// TIA Portal project "EEEB EMBU 4_V17" (V17)

(* hardware
DEVICE "ET 200SP station_1"  ET 200SP-Station
   slot 0: "Rack_0"  Rack  6ES5 710-8MAx1
   slot 1: "EEEB EMBU"  CPU 1510SP-1 PN  6ES7 510-1DJ01-0AB0  V2.6
   slot 2: "SLOT1"  DI 16x24VDC ST  6ES7 131-6BH01-0BA0  V0.0
      slot 1: "SLOT1"  DI 16x24VDC ST
   slot 3: "SLOT2"  DI 16x24VDC ST  6ES7 131-6BH01-0BA0  V0.0
      slot 1: "SLOT2"  DI 16x24VDC ST
   slot 4: "SLOT3"  DI 16x24VDC ST  6ES7 131-6BH01-0BA0  V0.0
      slot 1: "SLOT3"  DI 16x24VDC ST
   slot 5: "SLOT4"  DI 16x24VDC ST  6ES7 131-6BH01-0BA0  V0.0
      slot 1: "SLOT4"  DI 16x24VDC ST
   slot 6: "SLOT5"  DI 16x24VDC ST  6ES7 131-6BH01-0BA0  V0.0
      slot 1: "SLOT5"  DI 16x24VDC ST
   slot 7: "SLOT6"  DQ 16x24VDC/0.5A ST  6ES7 132-6BH01-0BA0  V0.0
      slot 1: "SLOT6"  DQ 16x24VDC/0.5A ST
   slot 8: "SLOT7"  DQ 16x24VDC/0.5A ST  6ES7 132-6BH01-0BA0  V0.0
      slot 1: "SLOT7"  DQ 16x24VDC/0.5A ST
   slot 9: "SLOT8"  AI 8xI 2-,4-wire BA  6ES7 134-6GF00-0AA1  V1.0
      slot 1: "SLOT8"  AI 8xI 2-,4-wire BA
   slot 10: "SLO9"  AI 8xI 2-,4-wire BA  6ES7 134-6GF00-0AA1  V1.0
      slot 1: "SLO9"  AI 8xI 2-,4-wire BA
   slot 11: "SLOT10"  AQ 4xU/I ST  6ES7 135-6HD00-0BA1  V1.1
      slot 1: "SLOT10"  AQ 4xU/I ST
   slot 12: "SLOT11"  AQ 4xU/I ST  6ES7 135-6HD00-0BA1  V1.1
      slot 1: "SLOT11"  AQ 4xU/I ST
   slot 13: "Server module_1"  Server module  6ES7 193-6PA00-0AA0  V1.1
      slot 1: "Server module_1"  Server module
   slot 127: "BA 2xRJ45"  BA 2xRJ45  6ES7 193-6AR00-0AA0  V0.0
      slot 32769: "Port_1"  6ES7 193-6AR00-0AA0
      slot 32770: "Port_2"  6ES7 193-6AR00-0AA0
DEVICE "HMI_1"  KTP700 Basic PN
   slot 0: "HMI_1"  KTP700 Basic PN  6AV2 123-2GB03-0AX0  15.1.0.0
   slot 1: "HMI_RT_1"  KTP700 Basic PN  6AV2 123-2GB03-0AX0  15.1.0.0
   slot 5: "HMI_1.IE_CP_1"  PROFINET Interface  15.0.1.0
      slot 1: "PROFINET Interface_1"  PROFINET Interface
         slot 1: "Port_1"  Port
*)

// ===== PLC "EEEB EMBU"  CPU 1510SP-1 PN =====

VAR_GLOBAL   // PLC tag table "Default tag table"
   "System_Byte" AT %MB1 : Byte;
   "FirstScan" AT %M1.0 : Bool;
   "DiagStatusUpdate" AT %M1.1 : Bool;
   "AlwaysTRUE" AT %M1.2 : Bool;
   "AlwaysFALSE" AT %M1.3 : Bool;
   "Clock_Byte" AT %MB0 : Byte;
   "Clock_10Hz" AT %M0.0 : Bool;
   "Clock_5Hz" AT %M0.1 : Bool;
   "Clock_2.5Hz" AT %M0.2 : Bool;
   "Clock_2Hz" AT %M0.3 : Bool;
   "Clock_1.25Hz" AT %M0.4 : Bool;
   "Clock_1Hz" AT %M0.5 : Bool;
   "Clock_0.625Hz" AT %M0.6 : Bool;
   "Clock_0.5Hz" AT %M0.7 : Bool;
   "Tag_3" AT %M50.0 : Bool;
   "bloqueio_provisorio" AT %M2.0 : Bool;
   "pause" AT %M2.1 : Bool;
   "bloqueio_provisorio_1" AT %M2.2 : Bool;
   "Tag_4" AT %M83.0 : Bool;
   "CON_MOD" AT %MW80 : Int;
   "INI" AT %M82.0 : Bool;
END_VAR

VAR_GLOBAL   // PLC tag table "IO"
   "PCM_EEE_EMER" AT %I0.0 : Bool;   // PCM-E-CF-01-04 BOTAO DE EMERGENCIA - ATUADO
   "PCM_EEE_K27" AT %I0.1 : Bool;   // PCM-E-CF-01-04 RELE DE PROTECAO FUNCAO 27 - ATUADO
   "PCM_EEE_DJL" AT %I0.2 : Bool;   // PCM-E-CF-01-04 DISJUNTOR GERAL STATUS - LIGADO
   "PCM_EEE_DJD" AT %I0.3 : Bool;   // PCM-E-CF-01-04 DISJUNTOR GERAL STATUS - DESLIGADO
   "PCM_EEE_DJYFAL" AT %I0.4 : Bool;   // PCM-E-CF-01-04 DISJUNTOR GERAL STATUS - FALHA
   "PCM_EEE_DJFG" AT %I0.5 : Bool;   // PCM-E-CF-01-04 FALHA GERAL ATUADO
   "PCM_EEE_TR01_KA3" AT %I0.6 : Bool;   // PCM-E-CF-01-04 TRANSFORMADOR -TR-01 ALARME TEMP 150°
   "PCM_EEE_TR01_KA4" AT %I0.7 : Bool;   // PCM-E-CF-01-04 TRANSFORMADOR -TR-01 ALARME TEMP 155°
   "PCM_EEE_TR01_KA5" AT %I1.0 : Bool;   // PCM-E-CF-01-04 TRANSFORMADOR -TR-01 FALHA PROTECAO
   "PCM_EEE_INTRU" AT %I1.1 : Bool;   // PCM-E-CF-01-04 INTRUSAO NO PAINEL (COLUNA 01~04)
   "MB_01_FF" AT %I1.2 : Bool;   // MB-01 FALTA DE FASE
   "MB_01_MMNT" AT %I1.3 : Bool;   // MB-01 MODO MANUTENCAO
   "MB_01_ML" AT %I1.4 : Bool;   // MB-01 MODO LOCAL
   "MB_01_MA" AT %I1.5 : Bool;   // MB-01 MODO AUTOMATICO
   "MB_01_MN" AT %I1.6 : Bool;   // MB-01 MODO NORMAL
   "MB_01_HMNT" AT %I1.7 : Bool;   // MB-01 HABILITA MANUTENCAO
   "MB_01_BL" AT %I2.0 : Bool;   // MB-01 BOMBA LIGADA
   "MB_01_DINV" AT %I2.1 : Bool;   // MB-01 DEFEITO NO INVERSOR
   "MB_01_DMB" AT %I2.2 : Bool;   // MB-01 DEFEITO NA BOMBA
   "MB_01_RST" AT %I2.3 : Bool;   // MB-01 RESET
   "MB_01_INTRU" AT %I2.4 : Bool;   // MB-01 INTRUSAO NO PAINEL
   "MB_01_EMER" AT %I2.5 : Bool;   // MB-01 EMERGENCIA
   "MB_02_FF" AT %I2.6 : Bool;   // MB-02 FALTA DE FASE
   "MB_02_MMNT" AT %I2.7 : Bool;   // MB-02 MODO MANUTENCAO
   "MB_02_ML" AT %I3.0 : Bool;   // MB-02 MODO LOCAL
   "MB_02_MA" AT %I3.1 : Bool;   // MB-02 MODO AUTOMATICO
   "MB_02_MN" AT %I3.2 : Bool;   // MB-02 MODO NORMAL
   "MB_02_HMNT" AT %I3.3 : Bool;   // MB-02 HABILITA MANUTENCAO
   "MB_02_BL" AT %I3.4 : Bool;   // MB-02 BOMBA LIGADA
   "MB_02_DINV" AT %I3.5 : Bool;   // MB-02 DEFEITO NO INVERSOR
   "MB_02_DMB" AT %I3.6 : Bool;   // MB-02 DEFEITO NA BOMBA
   "MB_02_RST" AT %I3.7 : Bool;   // MB-02 RESET
   "MB_02_INTRU" AT %I4.0 : Bool;   // MB-02 INTRUSAO NO PAINEL
   "MB_02_EMER" AT %I4.1 : Bool;   // MB-02 EMERGENCIA
   "MB_03_FF" AT %I4.2 : Bool;   // MB-03 FALTA DE FASE
   "MB_03_MMNT" AT %I4.3 : Bool;   // MB-03 MODO MANUTENCAO
   "MB_03_ML" AT %I4.4 : Bool;   // MB-03 MODO LOCAL
   "MB_03_MA" AT %I4.5 : Bool;   // MB-03 MODO AUTOMATICO
   "MB_03_MN" AT %I4.6 : Bool;   // MB-03 MODO NORMAL
   "MB_03_HMNT" AT %I4.7 : Bool;   // MB-03 HABILITA MANUTENCAO
   "MB_03_BL" AT %I5.0 : Bool;   // MB-03 BOMBA LIGADA
   "MB_03_DINV" AT %I5.1 : Bool;   // MB-03 DEFEITO NO INVERSOR
   "MB_03_DMB" AT %I5.2 : Bool;   // MB-03 DEFEITO NA BOMBA
   "MB_03_RST" AT %I5.3 : Bool;   // MB-03 RESET
   "MB_03_INTRU" AT %I5.4 : Bool;   // MB-03 INTRUSAO NO PAINEL
   "MB_03_EMER" AT %I5.5 : Bool;   // MB-03EMERGENCIA
   "MB_04_FF" AT %I5.6 : Bool;   // MB-04 FALTA DE FASE
   "MB_04_MMNT" AT %I5.7 : Bool;   // MB-04 MODO MANUTENCAO
   "MB_04_ML" AT %I6.0 : Bool;   // MB-04 MODO LOCAL
   "MB_04_MA" AT %I6.1 : Bool;   // MB-04 MODO AUTOMATICO
   "MB_04_MN" AT %I6.2 : Bool;   // MB-04 MODO NORMAL
   "MB_04_HMNT" AT %I6.3 : Bool;   // MB-04 HABILITA MANUTENCAO
   "MB_04_BL" AT %I6.4 : Bool;   // MB-04 BOMBA LIGADA
   "MB_04_DINV" AT %I6.5 : Bool;   // MB-04 DEFEITO NO INVERSOR
   "MB_04_DMB" AT %I6.6 : Bool;   // MB-04 DEFEITO NA BOMBA
   "MB_04_RST" AT %I6.7 : Bool;   // MB-04 RESET
   "MB_04_INTRU" AT %I7.0 : Bool;   // MB-04 INTRUSAO NO PAINEL
   "MB_04_EMER" AT %I7.1 : Bool;   // MB-04 EMERGENCIA
   "QGBT_EMER" AT %I7.2 : Bool;   // QGBT-AUX-01 BOTAO DE EMERGENCIA ATUADO
   "QGBT_K27" AT %I7.3 : Bool;   // QGBT-AUX-01 RELE DE PROTECAO FUNCAO 27/59 ATUADO
   "QGBT_DISJ_LIG" AT %I7.4 : Bool;   // QGBT-AUX-01 DISJUNTOR GERAL STATUS - LIGADO
   "QGBT_DISJ_DESLIG" AT %I7.5 : Bool;   // QGBT-AUX-01 DISJUNTOR GERAL STATUS - DESLIGADO
   "QGBT_DISJ_YFAL" AT %I7.6 : Bool;   // QGBT-AUX-01 DISJUNTOR GERAL FALHA - TRIP
   "QGBT_INTRU" AT %I7.7 : Bool;   // QGBT-AUX-01 INTRUSAO NO PAINEL
   "KI165" AT %I8.0 : Bool;   // RESERVA
   "KI166" AT %I8.1 : Bool;   // RESERVA
   "KI167" AT %I8.2 : Bool;   // RESERVA
   "KI168" AT %I8.3 : Bool;   // RESERVA
   "KI169" AT %I8.4 : Bool;   // RESERVA
   "KI170" AT %I8.5 : Bool;   // RESERVA
   "KI171" AT %I8.6 : Bool;   // RESERVA
   "KI172" AT %I8.7 : Bool;   // RESERVA
   "LSL_001" AT %I9.0 : Bool;   // CHAVE DE NIVEL -LSL-001
   "LSH_001" AT %I9.1 : Bool;   // CHAVE DE NIVEL -LSH-001
   "LSL_002" AT %I9.2 : Bool;   // CHAVE DE NIVEL -LSL-002
   "LSH_002" AT %I9.3 : Bool;   // CHAVE DE NIVEL -LSH-002
   "PCE_EEE_INTRU" AT %I9.4 : Bool;   // INTRUSAO NO PAINEL
   "PCE_EEE_UPS_ALM" AT %I9.5 : Bool;   // UPS EM ALARME FALHA NA BATERIA
   "PCE_EEE_UPS_FE" AT %I9.6 : Bool;   // UPS EM OPERACAO FALTA DE ENERGIA
   "PCE_EEE_UPS_CHAR" AT %I9.7 : Bool;   // UPS EM ALARME BATERIA CARREGADA
   "MB_01_SH" AT %Q0.0 : Bool;   // MB-01 SOLICITACAO HIDRAULICA
   "MB_01_PH" AT %Q0.1 : Bool;   // MB-01 PROTECAO HIDRAULICA
   "MB_01_INTV" AT %Q0.2 : Bool;   // MB-01 INTERVALO (COM)
   "MB_01_RR" AT %Q0.3 : Bool;   // MB-01 RESET REMOTO
   "MB_01_INTVS" AT %Q0.4 : Bool;   // MB-01 INTERVALO SINAL
   "MB_02_SH" AT %Q0.5 : Bool;   // MB-02 SOLICITACAO HIDRAULICA
   "MB_02_PH" AT %Q0.6 : Bool;   // MB-02 PROTECAO HIDRAULICA
   "MB_02_INTV" AT %Q0.7 : Bool;   // MB-02 INTERVALO (COM)
   "MB_02_RR" AT %Q1.0 : Bool;   // MB-02 RESET REMOTO
   "MB_02_INTVS" AT %Q1.1 : Bool;   // MB-02 INTERVALO SINAL
   "MB_03_SH" AT %Q1.2 : Bool;   // MB-03 SOLICITACAO HIDRAULICA
   "MB_03_PH" AT %Q1.3 : Bool;   // MB-03 PROTECAO HIDRAULICA
   "MB_03_INTV" AT %Q1.4 : Bool;   // MB-03 INTERVALO (COM)
   "MB_03_RR" AT %Q1.5 : Bool;   // MB-03 RESET REMOTO
   "MB_03_INTVS" AT %Q1.6 : Bool;   // MB-03 INTERVALO SINAL
   "MB_04_SH" AT %Q1.7 : Bool;   // MB-04 SOLICITACAO HIDRAULICA
   "LIT_001" AT %IW10 : Int;   // -LIT-001 TRANSMISSOR DE NIVEL TANQUE (TIPO RADAR)
   "MB_01_REF_VEL" AT %IW12 : Int;   // REFERENCIA DE VELOCIDADE INVERSOR DE FREQUENCIA BOMBA 01
   "MB_02_REF_VEL" AT %IW14 : Int;   // REFERENCIA DE VELOCIDADE INVERSOR DE FREQUENCIA BOMBA 02
   "MB_03_REF_VEL" AT %IW16 : Int;   // REFERENCIA DE VELOCIDADE INVERSOR DE FREQUENCIA BOMBA 03
   "MB_04_REF_VEL" AT %IW18 : Int;   // REFERENCIA DE VELOCIDADE INVERSOR DE FREQUENCIA BOMBA 04
   "FB6" AT %IW20 : Int;   // RESERVA
   "FB7" AT %IW22 : Int;   // RESERVA
   "FB8" AT %IW24 : Int;   // RESERVA
   "FB9" AT %IW26 : Int;   // RESERVA
   "FB10" AT %IW28 : Int;   // RESERVA
   "FB11" AT %IW30 : Int;   // RESERVA
   "FB12" AT %IW32 : Int;   // RESERVA
   "FB13" AT %IW34 : Int;   // RESERVA
   "FB14" AT %IW36 : Int;   // RESERVA
   "FB15" AT %IW38 : Int;   // RESERVA
   "FB16" AT %IW40 : Int;   // RESERVA
   "MB_01_VEL" AT %QW4 : Int;   // SETPOINT INVERSOR DE FREQUENCIA BOMBA 01
   "MB_02_VEL" AT %QW6 : Int;   // SETPOINT INVERSOR DE FREQUENCIA BOMBA 02
   "MB_03_VEL" AT %QW8 : Int;   // SETPOINT INVERSOR DE FREQUENCIA BOMBA 03
   "MB_04_VEL" AT %QW10 : Int;   // SETPOINT INVERSOR DE FREQUENCIA BOMBA 04
   "F25" AT %QW12 : Int;   // RESERVA
   "F26" AT %QW14 : Int;   // RESERVA
   "F27" AT %QW16 : Int;   // RESERVA
   "F28" AT %QW18 : Int;   // RESERVA
   "MB_04_PH" AT %Q2.0 : Bool;   // MB-04 PROTECAO HIDRAULICA
   "MB_04_INTV" AT %Q2.1 : Bool;   // MB-04 INTERVALO (COM)
   "MB_04_RR" AT %Q2.2 : Bool;   // MB-04 RESET REMOTO
   "MB_04_INTVS" AT %Q2.3 : Bool;   // MB-04 INTERVALO SINAL
   "KO21" AT %Q2.4 : Bool;   // RESERVA
   "KO22" AT %Q2.5 : Bool;   // RESERVA
   "KO23" AT %Q2.6 : Bool;   // RESERVA
   "KO24" AT %Q2.7 : Bool;   // RESERVA
   "KO25" AT %Q3.0 : Bool;   // RESERVA
   "KO26" AT %Q3.1 : Bool;   // RESERVA
   "KO27" AT %Q3.2 : Bool;   // RESERVA
   "KO28" AT %Q3.3 : Bool;   // RESERVA
   "KO29" AT %Q3.4 : Bool;   // RESERVA
   "KO30" AT %Q3.5 : Bool;   // RESERVA
   "KO31" AT %Q3.6 : Bool;   // RESERVA
   "KO32" AT %Q3.7 : Bool;   // RESERVA
END_VAR

VAR_GLOBAL   // PLC tag table "ALARMES"
   "ALM0" AT %MW100 : Word;   // ALARMES MB-01
   "ALM2" AT %MW102 : Word;   // ALARMES MB-02
   "ALM4" AT %MW104 : Word;   // ALARMES MB-03
   "ALM6" AT %MW106 : Word;   // ALARMES MB-04
   "ALM8" AT %MW108 : Word;   // ALARMES LIT_001
   "ALM10" AT %MW110 : Word;   // ALARMES PCM-EEE
   "ALM12" AT %MW112 : Word;   // ALARMES QGBT
   "ALM14" AT %MW114 : Word;   // ALARMES CHAVE DE NIVEL
   "ALM16" AT %MW116 : Word;   // ALARMES PCE-EEE
END_VAR

DATA_BLOCK "DIVERSOS"   // DB1
{ S7_Optimized_Access := 'TRUE' }
VERSION : 0.1
   VAR
      T1S : Bool;   // PULSO A CADA 1 SEGUNDO
      AUX_T1S : Bool;   // PULSO A CADA 1 SEGUNDO
      QTDE_PULSO : DInt := 200;
      ForcePulso : Bool;
      N_L00P : Int;
      Aux_N_LOOP : Int;
      Looping : Int := 0;
      TMR : Array[0..10] of IEC_TIMER;
      P1S : Bool;   // Pulso de 1 segundo
      "MB-01-SP" : Bool;   // Solicitação partida de bomba
      "MB-02-SP" : Bool;   // Solicitação partida de bomba
      "MB-03-SP" : Bool;   // Solicitação partida de bomba
      "MB-04-SP" : Bool;   // Solicitação partida de bomba
   END_VAR
BEGIN
END_DATA_BLOCK

DATA_BLOCK "INTPRO_DB"   // DB2
{ S7_Optimized_Access := 'TRUE' }
VERSION : 0.1
// stored: InstanceOfName INTPRO
"INTPRO"
BEGIN
END_DATA_BLOCK

DATA_BLOCK "LOOP_DB"   // DB3
{ S7_Optimized_Access := 'TRUE' }
VERSION : 0.1
// stored: InstanceOfName LOOP
"LOOP"
BEGIN
END_DATA_BLOCK

DATA_BLOCK "ROD4_DB"   // DB9
{ S7_Optimized_Access := 'FALSE' }
VERSION : 0.1
// stored: InstanceOfName ROD4
"ROD4"
BEGIN
END_DATA_BLOCK

DATA_BLOCK "ANALOGICOS_DB"   // DB101
{ S7_Optimized_Access := 'TRUE' }
VERSION : 0.1
// stored: InstanceOfName ANALOGICOS
"ANALOGICOS"
BEGIN
END_DATA_BLOCK

DATA_BLOCK "MODBUS_DB"   // DB102
{ S7_Optimized_Access := 'TRUE' }
VERSION : 0.1
// stored: InstanceOfName MODBUS
"MODBUS"
BEGIN
END_DATA_BLOCK

DATA_BLOCK "Digitais"   // DB300
{ S7_Optimized_Access := 'FALSE' }
VERSION : 0.1
   VAR
      "MB-01-YSH" : Bool;   // Elevatoria principal 1 ligado
      "MB-01-YR" : Bool;   // Elevatoria principal 1 remoto
      "MB-01-YF" : Bool;   // Elevatoria principal 1 falha
      "MB-01-YFF" : Bool;   // Elevatoria principal 1 falta de fase
      "MB-01-MM" : Bool;   // Elevatoria principal 1 modo manutenção
      "MB-01-MA" : Bool;   // Elevatoria principal 1 modo automatico
      "MB-01-EMER" : Bool;   // Elevatoria principal 1 emergencia
      "MB-01-MN" : Bool;   // Elevatoria principal 1 modo normal
      "MB-01-ML" : Bool;   // Elevatoria principal 1 modo local
      "MB-01-YFI" : Bool;   // Elevatoria principal 1 com falha no inversor
      "MB-01-YFA" : Bool;   // Elevatoria principal 1 com falha no acionamento
      "MB-01-YPTA" : Bool;   // Elevatoria principal 1 com proteção térmica atuada
      "MB-01-HM" : Bool;   // Elevatoria principal 1 habilita manutenção
      "MB-01-RST" : Bool;   // Elevatoria principal 1 reset
      "MB-01-INTRU" : Bool;   // Elevatoria principal 1 intrusão no painel
      "MB-01-YFB" : Bool;   // Elevatoria principal 1 defeito na bomba
      "MB-02-YSH" : Bool;   // Elevatoria principal 2 ligado
      "MB-02-YR" : Bool;   // Elevatoria principal 2 remoto
      "MB-02-YF" : Bool;   // Elevatoria principal 2 falha
      "MB-02-YFF" : Bool;   // Elevatoria principal 2 falta de fase
      "MB-02-MM" : Bool;   // Elevatoria principal 2 modo manutenção
      "MB-02-MA" : Bool;   // Elevatoria principal 2 modo automatico
      "MB-02-EMER" : Bool;   // Elevatoria principal 2 emergencia
      "MB-02-MN" : Bool;   // Elevatoria principal 2 modo normal
      "MB-02-ML" : Bool;   // Elevatoria principal 2 modo local
      "MB-02-YFI" : Bool;   // Elevatoria principal 2 com falha no inversor
      "MB-02-YFA" : Bool;   // Elevatoria principal 2 com falha no acionamento
      "MB-02-YPTA" : Bool;   // Elevatoria principal 2 com proteção térmica atuada
      "MB-02-HM" : Bool;   // Elevatoria principal 2 habilita manutenção
      "MB-02-RST" : Bool;   // Elevatoria principal 2 reset
      "MB-02-INTRU" : Bool;   // Elevatoria principal 2 intrusão no painel
      "MB-02-YFB" : Bool;   // Elevatoria principal 2 defeito na bomba
      "MB-03-YSH" : Bool;   // Elevatoria principal 3 ligado
      "MB-03-YR" : Bool;   // Elevatoria principal 3 remoto
      "MB-03-YF" : Bool;   // Elevatoria principal 3 falha
      "MB-03-YFF" : Bool;   // Elevatoria principal 3 falta de fase
      "MB-03-MM" : Bool;   // Elevatoria principal 3 modo manutenção
      "MB-03-MA" : Bool;   // Elevatoria principal 3 modo automatico
      "MB-03-EMER" : Bool;   // Elevatoria principal 3 emergencia
      "MB-03-MN" : Bool;   // Elevatoria principal 3 modo normal
      "MB-03-ML" : Bool;   // Elevatoria principal 3 modo local
      "MB-03-YFI" : Bool;   // Elevatoria principal 3 com falha no inversor
      "MB-03-YFA" : Bool;   // Elevatoria principal 3 com falha no acionamento
      "MB-03-YPTA" : Bool;   // Elevatoria principal 3 com proteção térmica atuada
      "MB-03-HM" : Bool;   // Elevatoria principal 3 habilita manutenção
      "MB-03-RST" : Bool;   // Elevatoria principal 3 reset
      "MB-03-INTRU" : Bool;   // Elevatoria principal 3 intrusão no painel
      "MB-03-YFB" : Bool;   // Elevatoria principal 3 defeito na bomba
      "MB-04-YSH" : Bool;   // Elevatoria principal 4 ligado
      "MB-04-YR" : Bool;   // Elevatoria principal 4 remoto
      "MB-04-YF" : Bool;   // Elevatoria principal 4 falha
      "MB-04-YFF" : Bool;   // Elevatoria principal 4 falta de fase
      "MB-04-MM" : Bool;   // Elevatoria principal 4 modo manutenção
      "MB-04-MA" : Bool;   // Elevatoria principal 4 modo automatico
      "MB-04-EMER" : Bool;   // Elevatoria principal 4 emergencia
      "MB-04-MN" : Bool;   // Elevatoria principal 4 modo normal
      "MB-04-ML" : Bool;   // Elevatoria principal 4 modo local
      "MB-04-YFI" : Bool;   // Elevatoria principal 4 com falha no inversor
      "MB-04-YFA" : Bool;   // Elevatoria principal 4 com falha no acionamento
      "MB-04-YPTA" : Bool;   // Elevatoria principal 4 com proteção térmica atuada
      "MB-04-HM" : Bool;   // Elevatoria principal 4 habilita manutenção
      "MB-04-RST" : Bool;   // Elevatoria principal 4 reset
      "MB-04-INTRU" : Bool;   // Elevatoria principal 4 intrusão no painel
      "MB-04-YFB" : Bool;   // Elevatoria principal 4 defeito na bomba
      "LIT_001-AL8" : Bool;   // Disponível para alarme
      "LIT_001-AL9" : Bool;   // Disponível para alarme
      "LIT_001-AL10" : Bool;   // Disponível para alarme
      "LIT_001-AL11" : Bool;   // Disponível para alarme
      "LIT_001-AL12" : Bool;   // Disponível para alarme
      "LIT_001-AL13" : Bool;   // Disponível para alarme
      "LIT_001-AL14" : Bool;   // Disponível para alarme
      "LIT_001-AL15" : Bool;   // Disponível para alarme
      "LIT_001-YHH" : Bool;   // Alarme de nível muito alto do tanque
      "LIT_001-YH" : Bool;   // Alarme de nível alto do tanque
      "LIT_001-YL" : Bool;   // Alarme de nível baixo do tanque
      "LIT_001-YLL" : Bool;   // Alarme de nível muito baixo do tanque
      "LIT_001-YFS" : Bool;   // Transmissor de nível do tanque com falha de sinal
      "LIT_001-AL5" : Bool;   // Disponível para alarme
      "LIT_001-AL6" : Bool;   // Disponível para alarme
      "LIT_001-AL7" : Bool;   // Disponível para alarme
      PCM_EEE_EMER : Bool;   // PCM-E-CF-01-04 BOTAO DE EMERGENCIA - ATUADO
      PCM_EEE_K27 : Bool;   // PCM-E-CF-01-04 RELE DE PROTECAO FUNCAO 27 - ATUADO
      PCM_EEE_DISJ_LIG : Bool;   // PCM-E-CF-01-04 DISJUNTOR GERAL STATUS - LIGADO
      PCM_EEE_DISJ_DESLIG : Bool;   // PCM-E-CF-01-04 DISJUNTOR GERAL STATUS - DESLIGADO
      PCM_EEE_DISJ_YFAL : Bool;   // PCM-E-CF-01-04 DISJUNTOR GERAL STATUS - FALHA
      PCM_EEE_DISJ_FAL_GR : Bool;   // PCM-E-CF-01-04 FALHA GERAL ATUADO
      PCM_EEE_TR01_KA3 : Bool;   // PCM-E-CF-01-04 TRANSFORMADOR -TR-01 ALARME TEMP 150°
      PCM_EEE_TR01_KA4 : Bool;   // PCM-E-CF-01-04 TRANSFORMADOR -TR-01 ALARME TEMP 155°
      PCM_EEE_TR01_KA5 : Bool;   // PCM-E-CF-01-04 TRANSFORMADOR -TR-01 FALHA PROTECAO
      PCM_EEE_INTRU : Bool;   // PCM-E-CF-01-04 INTRUSAO NO PAINEL (COLUNA 01~04)
      PCM_EEE_RSERVA_0 : Bool;   // PCM-E-CF-01-04 BIT RESERVA DA WORD
      PCM_EEE_RSERVA_1 : Bool;   // PCM-E-CF-01-04 BIT RESERVA DA WORD
      PCM_EEE_RSERVA_2 : Bool;   // PCM-E-CF-01-04 BIT RESERVA DA WORD
      PCM_EEE_RSERVA_3 : Bool;   // PCM-E-CF-01-04 BIT RESERVA DA WORD
      PCM_EEE_RSERVA_4 : Bool;   // PCM-E-CF-01-04 BIT RESERVA DA WORD
      PCM_EEE_RSERVA_5 : Bool;   // PCM-E-CF-01-04 BIT RESERVA DA WORD
      QGBT_EMER : Bool;   // QGBT-AUX-01 BOTAO DE EMERGENCIA ATUADO
      QGBT_K27 : Bool;   // QGBT-AUX-01 RELE DE PROTECAO FUNCAO 27/59 ATUADO
      QGBT_DJL : Bool;   // QGBT-AUX-01 DISJUNTOR GERAL STATUS - LIGADO
      QGBT_DJD : Bool;   // QGBT-AUX-01 DISJUNTOR GERAL STATUS - DESLIGADO
      QGBT_DJYFAL : Bool;   // QGBT-AUX-01 DISJUNTOR GERAL FALHA - TRIP
      QGBT_INTRU : Bool;   // QGBT-AUX-01 INTRUSAO NO PAINEL
      QGBT_RESERVA_0 : Bool;   // QGBT-AUX-01 BIT RESERVA DA WORD
      QGBT_RESERVA_1 : Bool;   // QGBT-AUX-01 BIT RESERVA DA WORD
      QGBT_RESERVA_2 : Bool;   // QGBT-AUX-01 BIT RESERVA DA WORD
      QGBT_RESERVA_3 : Bool;   // QGBT-AUX-01 BIT RESERVA DA WORD
      QGBT_RESERVA_4 : Bool;   // QGBT-AUX-01 BIT RESERVA DA WORD
      QGBT_RESERVA_5 : Bool;   // QGBT-AUX-01 BIT RESERVA DA WORD
      QGBT_RESERVA_6 : Bool;   // QGBT-AUX-01 BIT RESERVA DA WORD
      QGBT_RESERVA_7 : Bool;   // QGBT-AUX-01 BIT RESERVA DA WORD
      QGBT_RESERVA_8 : Bool;   // QGBT-AUX-01 BIT RESERVA DA WORD
      QGBT_RESERVA_9 : Bool;   // QGBT-AUX-01 BIT RESERVA DA WORD
      LSL_001 : Bool;   // CHAVE DE NIVEL -LSL-001
      LSH_001 : Bool;   // CHAVE DE NIVEL -LSH-001
      LSL_002 : Bool;   // CHAVE DE NIVEL -LSL-002
      LSH_002 : Bool;   // CHAVE DE NIVEL -LSH-002
      LS_RESERVA_0 : Bool;   // CHAVE DE NIVEL - LS BIT RESERVA DA WORD
      LS_RESERVA_1 : Bool;   // CHAVE DE NIVEL - LS BIT RESERVA DA WORD
      LS_RESERVA_2 : Bool;   // CHAVE DE NIVEL - LS BIT RESERVA DA WORD
      LS_RESERVA_3 : Bool;   // CHAVE DE NIVEL - LS BIT RESERVA DA WORD
      LS_RESERVA_4 : Bool;   // CHAVE DE NIVEL - LS BIT RESERVA DA WORD
      LS_RESERVA_5 : Bool;   // CHAVE DE NIVEL - LS BIT RESERVA DA WORD
      LS_RESERVA_6 : Bool;   // CHAVE DE NIVEL - LS BIT RESERVA DA WORD
      LS_RESERVA_7 : Bool;   // CHAVE DE NIVEL - LS BIT RESERVA DA WORD
      LS_RESERVA_8 : Bool;   // CHAVE DE NIVEL - LS BIT RESERVA DA WORD
      LS_RESERVA_9 : Bool;   // CHAVE DE NIVEL - LS BIT RESERVA DA WORD
      LS_RESERVA_10 : Bool;   // CHAVE DE NIVEL - LS BIT RESERVA DA WORD
      LS_RESERVA_11 : Bool;   // CHAVE DE NIVEL - LS BIT RESERVA DA WORD
      PCE_EEE_INTRU : Bool;   // INTRUSAO NO PAINEL
      PCE_EEE_UPS_ALM : Bool;   // UPS EM ALARME FALHA NA BATERIA
      PCE_EEE_UPS_FE : Bool;   // UPS EM OPERACAO FALTA DE ENERGIA
      PCE_EEE_UPS_CHAR : Bool;   // UPS EM ALARME BATERIA CARREGADA
      "PCM-E-CF-01-P100-YFC" : Bool;   // Falha de comunicação com medidor do PCM-E-CF-01
      "QGBT-AUX-01-P100-YFC" : Bool;   // Falha de comunicação com medidor do PCM-E-CF-02
   END_VAR
BEGIN
END_DATA_BLOCK

DATA_BLOCK "ALARMES"   // DB301
{ S7_Optimized_Access := 'TRUE' }
VERSION : 0.1
   VAR
      "CCM-02-EA-P100-YFC" : Bool;   // Falha de comunicação com medidor do CCM1
      "CCM-02-EB-P100-YFC" : Bool;   // Falha de comunicação com medidor do CCM2
      "LIT_001-YHH" : Bool;   // Alarme de nível muito alto do tanque água bruta
      "LIT_001-YH" : Bool;   // Alarme de nível alto do tanque água bruta
      "LIT_001-YL" : Bool;   // Alarme de nível baixo do tanque água bruta
      "LIT_001-YLL" : Bool;   // Alarme de nível muito baixo do tanque água bruta
      "LIT_001-YFS" : Bool;   // Transmissor de nível do tanque água bruta com falha de sinal
      "LIT_001-YHHH" : Bool;   // Alarme de nível muito alto - desliga CAB e lavagem peneira
      "CAB-PT-015-YH" : Bool;
      "CAB-PT-015-YFS" : Bool;
      "MB-03-YIP" : Bool;   // MB-03 com intervalo entre partidas
      "MB-02-YIP" : Bool;   // MB-02 com intervalo entre partidas
      "MB-01-YIP" : Bool;   // MB-01 com intervalo entre partidas
   END_VAR
BEGIN
END_DATA_BLOCK

DATA_BLOCK "STATUS"   // DB302
{ S7_Optimized_Access := 'FALSE' }
VERSION : 0.1
   VAR
      "SO-203-06A-YI" : Bool;   // Soprador tanque de aeração intertravado
      "SO-203-06B-YI" : Bool;   // Soprador tanque de aeração intertravado
      "SO-203-06C-YI" : Bool;   // Soprador tanque de aeração intertravado
      "SO-203-06D-YI" : Bool;   // Soprador tanque de aeração intertravado
      "SO-203-06E-YI" : Bool;   // Soprador tanque de aeração intertravado
      "SO-203-06F-YI" : Bool;   // Soprador tanque de aeração intertravado
      "MB-01-YSP" : Bool;   // MB-01 selecionada como principal
      "MB-02-YSP" : Bool;   // MB-02 selecionada como principal
      "MB-04-YSP" : Bool;   // MB-03 selecionada como principal
      "MB-03-YSP" : Bool;   // MB-03 selecionada como principal
      "MB-01-YC1" : Bool;   // MB-01 selecionada como complementar 1
      "MB-02-YC1" : Bool;   // MB-02 selecionada como complementar 1
      "MB-04-YC1" : Bool;   // MB-03 selecionada como complementar 1
      "MB-03-YC1" : Bool;   // MB-03 selecionada como complementar 1
      "MB-01-YC2" : Bool;   // MB-01 selecionada como complementar 2
      "MB-02-YC2" : Bool;   // MB-02 selecionada como complementar 2
      "MB-04-YC2" : Bool;   // MB-03 selecionada como complementar 2
      "MB-03-YC2" : Bool;   // MB-03 selecionada como complementar 2
      "MB-01-YC3" : Bool;   // MB-01 selecionada como complementar 3
      "MB-02-YC3" : Bool;   // MB-02 selecionada como complementar 3
      "MB-04-YC3" : Bool;   // MB-03 selecionada como complementar 3
      "MB-03-YC3" : Bool;   // MB-03 selecionada como complementar 3
   END_VAR
BEGIN
END_DATA_BLOCK

DATA_BLOCK "COMANDOS"   // DB303
{ S7_Optimized_Access := 'FALSE' }
VERSION : 0.1
   VAR
      "MB-01-HS9" : Bool := false;   // Comando disponível
      "MB-01-HS10" : Bool := false;   // Comando disponível
      "MB-01-HS11" : Bool;   // Comando disponível
      "MB-01-HS12" : Bool;   // Comando disponível
      "MB-01-HS13" : Bool;   // Comando disponível
      "MB-01-HS14" : Bool;   // Comando disponível
      "MB-01-HS15" : Bool;   // Comando disponível
      "MB-01-HS16" : Bool;   // Comando disponível
      "MB-01-HS1" : Bool := true;   // Comando manual/automático
      "MB-01-HS2" : Bool := false;   // Comando liga
      "MB-01-HS3" : Bool := false;   // Comando desliga
      "MB-01-HS4" : Bool := false;   // Comando reset falha
      "MB-01-HS5" : Bool := false;   // Comando reset tempo de operação
      "MB-01-HS6" : Bool;
      "MB-01-HS7" : Bool := false;   // Comando habilita bloqueio
      "MB-01-HS8" : Bool := false;   // Comando disponível
      "MB-02-HS9" : Bool := false;   // Comando disponível
      "MB-02-HS10" : Bool := false;   // Comando disponível
      "MB-02-HS11" : Bool;   // Comando disponível
      "MB-02-HS12" : Bool;   // Comando disponível
      "MB-02-HS13" : Bool;   // Comando disponível
      "MB-02-HS14" : Bool;   // Comando disponível
      "MB-02-HS15" : Bool;   // Comando disponível
      "MB-02-HS16" : Bool;   // Comando disponível
      "MB-02-HS1" : Bool := true;   // Comando manual/automático
      "MB-02-HS2" : Bool := false;   // Comando liga
      "MB-02-HS3" : Bool := false;   // Comando desliga
      "MB-02-HS4" : Bool := false;   // Comando reset falha
      "MB-02-HS5" : Bool := false;   // Comando reset tempo de operação
      "MB-02-HS6" : Bool;
      "MB-02-HS7" : Bool := false;   // Comando habilita bloqueio
      "MB-02-HS8" : Bool := false;   // Comando disponível
      "MB-03-HS9" : Bool := false;   // Comando disponível
      "MB-03-HS10" : Bool := false;   // Comando disponível
      "MB-03-HS11" : Bool;   // Comando disponível
      "MB-03-HS12" : Bool;   // Comando disponível
      "MB-03-HS13" : Bool;   // Comando disponível
      "MB-03-HS14" : Bool;   // Comando disponível
      "MB-03-HS15" : Bool;   // Comando disponível
      "MB-03-HS16" : Bool;   // Comando disponível
      "MB-03-HS1" : Bool := true;   // Comando manual/automático
      "MB-03-HS2" : Bool := false;   // Comando liga
      "MB-03-HS3" : Bool := false;   // Comando desliga
      "MB-03-HS4" : Bool := false;   // Comando reset falha
      "MB-03-HS5" : Bool := false;   // Comando reset tempo de operação
      "MB-03-HS6" : Bool;
      "MB-03-HS7" : Bool := false;   // Comando habilita bloqueio
      "MB-03-HS8" : Bool := false;   // Comando disponível
      "MB-04-HS9" : Bool := false;   // Comando disponível
      "MB-04-HS10" : Bool := false;   // Comando disponível
      "MB-04-HS11" : Bool;   // Comando disponível
      "MB-04-HS12" : Bool;   // Comando disponível
      "MB-04-HS13" : Bool;   // Comando disponível
      "MB-04-HS14" : Bool;   // Comando disponível
      "MB-04-HS15" : Bool;   // Comando disponível
      "MB-04-HS16" : Bool;   // Comando disponível
      "MB-04-HS1" : Bool := false;   // Comando manual/automático
      "MB-04-HS2" : Bool := false;   // Comando liga
      "MB-04-HS3" : Bool := false;   // Comando desliga
      "MB-04-HS4" : Bool := false;   // Comando reset falha
      "MB-04-HS5" : Bool := false;   // Comando reset tempo de operação
      "MB-04-HS6" : Bool;
      "MB-04-HS7" : Bool := false;   // Comando habilita bloqueio
      "MB-04-HS8" : Bool := false;   // Comando disponível
      "LIT_001-HS9" : Bool;   // Comando disponível
      "LIT_001-HS10" : Bool;   // Comando disponível
      "LIT_001-HS11" : Bool;   // Comando disponível
      "LIT_001-HS12" : Bool;   // Comando disponível
      "LIT_001-HS13" : Bool;   // Comando disponível
      "LIT_001-HS14" : Bool;   // Comando disponível
      "LIT_001-HS15" : Bool;   // Comando disponível
      "LIT_001-HS16" : Bool;   // Comando disponível
      "LIT_001-HSHH" : Bool;   // Inibe alarme muito alto montante peneira 1
      "LIT_001-HSH" : Bool;   // Inibe alarme nível alto montante peneira 1
      "LIT_001-HSL" : Bool;   // Inibe alarme nível baixo montante peneira 1
      "LIT_001-HSLL" : Bool;   // Inibe alarme nível muito baixo montante peneira 1
      "LIT_001-HSM" : Bool;   // Habilita valor manual para medidor
      "LIT_001-HS6" : Bool;   // Comando disponível
      "LIT_001-HS7" : Bool;   // Comando disponível
      "LIT_001-HS8" : Bool;   // Comando disponível
      "PID-TA3-HI" : Bool;   // Habilita integrall PID tanque de aeração
      "PID-EEEB-HD" : Bool;   // Habilita derivativo PID tanque de aeração
      "PID-EEEB-HP" : Bool;   // Habilita proporcional PID tanque de aeração
      "PID-EEEB-HI" : Bool;   // Habilita integrall PID tanque de aeração
      "PID-TA5-HD" : Bool;   // Habilita derivativo PID tanque de aeração
      "PID-TA5-HP" : Bool;   // Habilita proporcional PID tanque de aeração
      "PID-TA5-HI" : Bool;   // Habilita integrall PID tanque de aeração
      "PID-TA1-HM" : Bool;   // Habilita valor manual para saída
      "PID-TA1-HD" : Bool;   // Habilita derivativo PID tanque de aeração
      "PID-TA1-HP" : Bool;   // Habilita proporcional PID tanque de aeração
      "PID-TA1-HI" : Bool;   // Habilita integrall PID tanque de aeração
      "PID-TA2-HD" : Bool;   // Habilita derivativo PID tanque de aeração
      "PID-TA2-HP" : Bool;   // Habilita proporcional PID tanque de aeração
      "PID-TA2-HI" : Bool;   // Habilita integrall PID tanque de aeração
      "PID-TA3-HD" : Bool;   // Habilita derivativo PID tanque de aeração
      "PID-TA3-HP" : Bool;   // Habilita proporcional PID tanque de aeração
      "PID-TA2-HM" : Bool;   // Habilita valor manual para saída
      "PID-TA3-HM" : Bool;   // Habilita valor manual para saída
      "PID-EEEB-HM" : Bool;   // Habilita valor manual para saída
      "PID-TA5-HM" : Bool;   // Habilita valor manual para saída
   END_VAR
BEGIN
END_DATA_BLOCK

DATA_BLOCK "VARIAVEIS"   // DB304
{ S7_Optimized_Access := 'FALSE' }
VERSION : 0.1
   VAR
      "MB-01-YST" : Real;   // Frequência raspador de areia
      "MB-01-YIT" : Real;   // Corrente raspador de areia
      "MB-02-YIT" : Real;   // Corrente raspador de areia
      "MB-02-YST" : Real;   // Frequência raspador de areia
      "MB-03-YIT" : Real;   // Corrente raspador de areia
      "MB-03-YST" : Real;   // Frequência raspador de areia
      "MB-04-YIT" : Real;   // Corrente raspador de areia
      "MB-04-YST" : Real;   // Frequência raspador de areia
      LIT_001 : Real;   // Nível Tanque
      "LIT_001-P" : Real;   // Percentual Tanque
      "PCM-E-CF-01-04-P100-ETRS" : Real;   // Tensão entre fases R e S
      "PCM-E-CF-01-04-P100-ETST" : Real;   // Tensão entre fases S e T
      "PCM-E-CF-01-04-P100-ETTR" : Real;   // Tensão entre fases T e R
      "PCM-E-CF-01-04-P100-ITR" : Real;   // Corrente fase R
      "PCM-E-CF-01-04-P100-ITS" : Real;   // Corrente fase S
      "PCM-E-CF-01-04-P100-ITT" : Real;   // Corrente fase T
      "PCM-E-CF-01-04-P100-JPT" : Real;   // Potência ativa total
      "PCM-E-CF-01-04-P100-JQT" : Real;   // Potência reativa total
      "PCM-E-CF-01-04-P100-JST" : Real;   // Potência aparente total
      "PCM-E-CF-01-04-P100-FP" : Real;   // Fator de potência
      "QGBT-AUX-01-P100-ETRS" : Real;   // Tensão entre fases R e S
      "QGBT-AUX-01-P100-ETST" : Real;   // Tensão entre fases S e T
      "QGBT-AUX-01-P100-ETTR" : Real;   // Tensão entre fases T e R
      "QGBT-AUX-01-P100-ITR" : Real;   // Corrente fase R
      "QGBT-AUX-01-P100-ITS" : Real;   // Corrente fase S
      "QGBT-AUX-01-P100-ITT" : Real;   // Corrente fase T
      "QGBT-AUX-01-P100-JPT" : Real;   // Potência ativa total
      "QGBT-AUX-01-P100-JQT" : Real;   // Potência reativa total
      "QGBT-AUX-01-P100-JST" : Real;   // Potência aparente total
      "QGBT-AUX-01-P100-FP" : Real;   // Fator de potência
   END_VAR
BEGIN
END_DATA_BLOCK

DATA_BLOCK "SETPOINTS"   // DB305
{ S7_Optimized_Access := 'FALSE' }
VERSION : 0.1
   VAR
      "MB-01-SP" : Real := 60.0;   // Setpoint manual elevatoria principal
      "MB-02-SP" : Real := 0.0;   // Setpoint manual elevatoria principal
      "MB-03-SP" : Real := 60.0;   // Setpoint manual elevatoria principal
      "MB-04-SP" : Real := 60.0;   // Setpoint manual elevatoria principal
      "LIT_001-SPHH" : Real := 90.0;   // Setpoint muito alto elevatoria principal
      "LIT_001-SPH" : Real := 70.0;   // Setpoint nível alto elevatoria principal
      "LIT_001-SPL" : Real := 10.0;   // Setpoint nível baixo elevatoria principal
      "LIT_001-SPLL" : Real := 0.0;   // Setpoint nível muito baixo elevatoria principal
      "LIT_001-SPM" : Real := 48.0;   // Habilita valor manual para medidor
      "LIT_001-SPC" : Real := 0.0;   // Setpoint de controle tanque
      "LIT-001-P" : Real := 0.0;
      SP_NVL_MIN : Real := 1.0;   // setpoint nivel minimo do tanque para proteção hidraulica
      "MB-P-SP-DL" : Real := 2.0;   // Setpoint para desligar bomba Principal
      "MB-P-SP-L" : Real := 2.6;   // Setpoint para ligar bomba Principal
      "MB-C1-SP-DL" : Real := 2.35;   // Setpoint para desligar bomba complementar 1
      "MB-C1-SP-L" : Real := 2.9;   // Setpoint para ligar bomba complementar 1
      "MB-C2-SP-DL" : Real := 2.66;   // Setpoint para desligar bomba complementar 2
      "MB-C2-SP-L" : Real := 3.9;   // Setpoint para ligar bomba complementar 2
      "MB-C3-SP-DL" : Real := 0.0;   // Setpoint para desligar bomba complementar 3
      "MB-C3-SP-L" : Real := 0.0;   // Setpoint para ligar bomba complementar 3
   END_VAR
BEGIN
END_DATA_BLOCK

DATA_BLOCK "Totalizadores"   // DB306
{ S7_Optimized_Access := 'FALSE' }
VERSION : 0.1
   VAR
      "MB-01-SO" : Int;   // Segundos em operação elevatoria principal
      "MB-01-MO" : Int;   // Minutos em operação elevatoria principal
      "MB-01-HO" : Int;   // Horas em operação elevatoria principal
      "MB-02-SO" : Int;   // Segundos em operação elevatoria principal
      "MB-02-MO" : Int;   // Minutos em operação elevatoria principal
      "MB-02-HO" : Int;   // Horas em operação elevatoria principal
      "MB-03-SO" : Int;   // Segundos em operação elevatoria principal
      "MB-03-MO" : Int;   // Minutos em operação elevatoria principal
      "MB-03-HO" : Int;   // Horas em operação elevatoria principal
      "MB-04-SO" : Int;   // Segundos em operação elevatoria principal
      "MB-04-MO" : Int;   // Minutos em operação elevatoria principal
      "MB-04-HO" : Int;   // Horas em operação elevatoria principal
   END_VAR
BEGIN
END_DATA_BLOCK

DATA_BLOCK "PID"   // DB307
{ S7_Optimized_Access := 'FALSE' }
VERSION : 0.1
   VAR
      "PID-EEEB-D" : Real;   // Ajuste derivativo PID elevatória de esgoto bruto
      "PID-EEEB-P" : Real;   // Ajuste proporcional PID elevatória de esgoto bruto
      "PID-EEEB-I" : Real;   // Ajuste integral PID elevatória de esgoto bruto
      "PID-EEEB-MIN" : Real;   // Ajuste mínimo PID elevatória de esgoto bruto
      "PID-EEEB-MAX" : Real;   // Ajuste máximo PID elevatória de esgoto bruto
      "PID-EEEB-DB" : Real;   // Banda morta PID elevatória de esgoto bruto
      "PID-EEEB-SPM" : Real;   // Setpoint manual
      "VA-PID-EEEB" : Real;   // Variável atuada PID elevatória de esgoto bruto
      "PID-EEEB-VR" : Real;   // Valor Relativo do PID
      AUX_CALC : Array[0..10] of Real;
   END_VAR
BEGIN
END_DATA_BLOCK

DATA_BLOCK "PDIR_DB_MB-01"   // DB422
{ S7_Optimized_Access := 'FALSE' }
VERSION : 0.1
// stored: InstanceOfName PDIR
"PDIR"
BEGIN
END_DATA_BLOCK

DATA_BLOCK "PDIR_DB_MB-02"   // DB423
{ S7_Optimized_Access := 'FALSE' }
VERSION : 0.1
// stored: InstanceOfName PDIR
"PDIR"
BEGIN
END_DATA_BLOCK

DATA_BLOCK "PDIR_DB_MB-03"   // DB424
{ S7_Optimized_Access := 'FALSE' }
VERSION : 0.1
// stored: InstanceOfName PDIR
"PDIR"
BEGIN
END_DATA_BLOCK

DATA_BLOCK "PDIR_DB_MB-04"   // DB425
{ S7_Optimized_Access := 'FALSE' }
VERSION : 0.1
// stored: InstanceOfName PDIR
"PDIR"
BEGIN
END_DATA_BLOCK

DATA_BLOCK "Redes"   // DB500
{ S7_Optimized_Access := 'FALSE' }